(* Logix 5000 project; controller MV vendor 1 type 14 code 217 rev 31.11; software revision 31.00; part 16 of 53 *)
(* tags used below, declared in another part *)
   CWD : CHECKWORD_FLAGS;
   Dummy : BOOL;
   MC_B12 : INT[255];   // PX SWITCH Proxy switch flags f ile
   MC_B240 : INT[255];   // CH1 RN PMP Channel 1 return pum p drive flags
   MC_B241 : INT[255];   // CH2 RN PMP Channel 2 return pum p drive flags
   MC_B242 : INT[255];   // CH1 ROUTE Channel 1 route requ est flags
   MC_B243 : INT[255];   // CH2 ROUTE Channel 2 route requ est flags
   MC_B3 : INT[255];   // BINARY
   MC_bit_data_file_address : DINT;
   MC_bit_file_bit_offset : DINT;
   MC_bit_file_word_offset : DINT;
   MC_bit_offset : DINT;
   MC_bit_returned : BOOL;
   MC_CP1 : PlantItem;   // CP1
   MC_CP1_RawOutput : ALIAS FOR RIO_Rack_2:10:O.Data.14;   // MC_CP1
   MC_data_file_value_to_move : DINT;
   MC_from_data_file : DINT;
   MC_from_data_offset : DINT;
   MC_GBYV1 : PlantItem;   // GBYV1
   MC_GBYV1_RawOutput : ALIAS FOR RIO_Rack_2:8:O.Data.31;   // MC_GBYV1
   MC_N10 : INT[255];   // SETTINGS
   MC_N100 : INT[255];   // C1_PLC Channel 1 PLC data
   MC_N101 : INT[255];   // CH1 PC>PLC Channel 1 PC to PLC
   MC_N102 : INT[255];   // CH1 PROG Channel 1 CIP progra m
   MC_N103 : INT[255];   // CH1 ITEMS Chwd.nos.of items to be checked for Chan nel 1
   MC_N104 : INT[255];   // CH1 REPORT Channel 1 CIP report file
   MC_N108 : INT[255];   // CH1 VDATA Channel 1 CIP progra m validation data
   MC_N112 : INT[255];   // FVR DATA Data read from FV ro uting PLC
   MC_N113 : INT[255];   // MVR DATA Data read from MV ro uting PLC
   MC_N114 : INT[255];   // YP DATA
   MC_N120 : INT[255];   // C2 PLC Channel 2 PLC data
   MC_N121 : INT[255];   // CH2 PC>PLC Channel 2 PC to PLC
   MC_N122 : INT[255];   // CH2 PROG Channel 2 CIP progra m
   MC_N123 : INT[255];   // CH2 ITEMS Chwd.nos.of items to be checked for Chan nel 2
   MC_N124 : INT[255];   // CH2 REPORT Channel 2 CIP report file
   MC_N128 : INT[255];   // CH2 VDATA Channel 2 CIP progra m validation data
   MC_N160 : INT[255];   // P40 CHECK
   MC_N161 : INT[255];   // P41 CHECK
   MC_N162 : INT[255];   // P42 CHECK
   MC_N163 : INT[255];   // P43 CHECK
   MC_N164 : INT[255];   // P44 CHECK
   MC_N165 : INT[255];   // P45 CHECK
   MC_N166 : INT[255];   // P46 CHECK
   MC_N167 : INT[255];   // Original N File From SLC, No Description Available
   MC_N20 : INT[255];   // P1 PRESS Control block and da ta for P1 pressure P ID loop
   MC_N200 : INT[255];   // CHK_WORK Plant item fault che cking work area
   MC_N201 : INT[255];   // P1 CHECK CIP program 1 plant item check list
   MC_N202 : INT[255];   // P2 CHECK CIP program 2 plant item check list
   MC_N203 : INT[255];   // P3 CHECK CIP program 3 plant item check list
   MC_N204 : INT[255];   // P4 CHECK CIP program 4 plant item check list
   MC_N205 : INT[255];   // P5 CHECK CIP program 5 plant item check list
   MC_N206 : INT[255];   // P6 CHECK CIP program 6 plant item check list
   MC_N207 : INT[255];   // P7 CHECK CIP program 7 plant item check list
   MC_N208 : INT[255];   // P8 CHECK CIP program 8 plant item check list
   MC_N209 : INT[255];   // P9 CHECK CIP program 9 plant item check list
   MC_N21 : INT[255];   // P1 FLOW Control block and da ta for P1 flowrate P ID loop
   MC_N210 : INT[255];   // P10 CHECK CIP program 10 plant item check list
   MC_N211 : INT[255];   // P11 CHECK CIP program 11 plant item check list
   MC_N212 : INT[255];   // P12 CHECK CIP program 12 plant item check list
   MC_N213 : INT[255];   // P13 CHECK CIP program 13 plant item check list
   MC_N214 : INT[255];   // P14 CHECK CIP program 14 plant item check list
   MC_N215 : INT[255];   // P15 CHECK CIP program 15 plant item check list
   MC_N216 : INT[255];   // P16 CHECK CIP program 16 plant item check list
   MC_N217 : INT[255];   // P17 CHECK CIP program 17 plant item check list
   MC_N218 : INT[255];   // P18 CHECK CIP program 18 plant item check list
   MC_N219 : INT[255];   // P19 CHECK CIP program 19 plant item check list
   MC_N22 : INT[255];   // P2 PRESS Control block and da ta for P2 pressure P ID loop
   MC_N220 : INT[255];   // P20 CHECK CIP program 20 plant item check list
   MC_N221 : INT[255];   // P21 CHECK CIP program 21 plant item check list
   MC_N222 : INT[255];   // P22 CHECK CIP program 22 plant item check list
   MC_N223 : INT[255];   // P23 CHECK CIP program 23 plant item check list
   MC_N224 : INT[255];   // P24 CHECK CIP program 24 plant item check list
   MC_N225 : INT[255];   // P25 CHECK CIP program 25 plant item check list
   MC_N226 : INT[255];   // P26 CHECK CIP program 26 plant item check list
   MC_N227 : INT[255];   // P27 CHECK CIP program 27 plant item check list
   MC_N228 : INT[255];   // P28 CHECK CIP program 28 plant item check list
   MC_N229 : INT[255];   // P29 CHECK CIP program 29 plant item check list
   MC_N23 : INT[255];   // P2 FLOW Control block and da ta for P2 flowrate P ID loop
   MC_N230 : INT[255];   // P30 CHECK CIP program 30 plant item check list
   MC_N231 : INT[255];   // P31 CHECK CIP program 31 plant item check list
   MC_N232 : INT[255];   // P32 CHECK CIP program 32 plant item check list
   MC_N233 : INT[255];   // P33 CHECK CIP program 33 plant item check list
   MC_N234 : INT[255];   // P34 CHECK CIP program 34 plant item check list
   MC_N235 : INT[255];   // P35 CHECK CIP program 35 plant item check list
   MC_N236 : INT[255];   // P36 CHECK CIP program 36 plant item check list
   MC_N237 : INT[255];   // P37 CHECK CIP program 37 plant item check list
   MC_N238 : INT[255];   // P38 CHECK CIP program 38 plant item check list
   MC_N239 : INT[255];   // P39 CHECK CIP program 39 plant item check list
   MC_N245 : INT[255];   // CC_WORK Continuous checking program work area
   MC_N255 : INT[255];   // CHECKWORDS Plant item checkword s
   MC_N7 : INT[255];   // INTEGER
   MC_N80 : INT[255];   // SRV1_PLC Detergent tank 1 ser vice PLC data
   MC_N81 : INT[255];   // SV1_PC Detergent tank 1 ser vice PC to PLC data
   MC_N82 : INT[255];   // SV1 ITEMS Chwd.nos.of items to be checked for DT1 service
   MC_N90 : INT[255];   // SV2_PLC Detergent tank 2 ser vice PLC data
   MC_N91 : INT[255];   // SV2_PC Detergent tank 2 ser vice PC to PLC data
   MC_N92 : INT[255];   // SV2 ITEMS Chwd.nos.of items to be checked for DT2 service
   MC_SP_V12TO17 : PlantItem;   // SP_V12TO17
   MC_SP_V12TO17_RawOutput : ALIAS FOR RIO_Rack_2:10:O.Data.17;   // MC_SP_V12TO17
(* MC_Common, continued *)

ROUTINE MC_Digital_Outputs   (* ladder *)
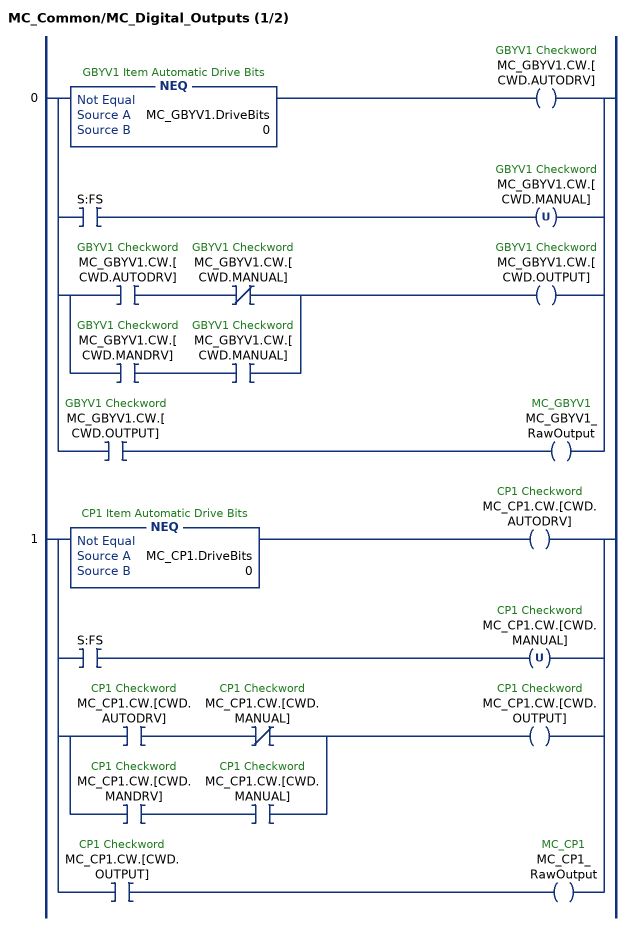
   0: [NEQ(MC_GBYV1.DriveBits,0) OTE(MC_GBYV1.CW.[CWD.AUTODRV]) ,XIC(S:FS) OTU(MC_GBYV1.CW.[CWD.MANUAL]) ,[XIC(MC_GBYV1.CW.[CWD.AUTODRV]) XIO(MC_GBYV1.CW.[CWD.MANUAL]) ,XIC(MC_GBYV1.CW.[CWD.MANDRV]) XIC(MC_GBYV1.CW.[CWD.MANUAL]) ] OTE(MC_GBYV1.CW.[CWD.OUTPUT]) ,XIC(MC_GBYV1.CW.[CWD.OUTPUT]) OTE(MC_GBYV1_RawOutput) ];
   1: [NEQ(MC_CP1.DriveBits,0) OTE(MC_CP1.CW.[CWD.AUTODRV]) ,XIC(S:FS) OTU(MC_CP1.CW.[CWD.MANUAL]) ,[XIC(MC_CP1.CW.[CWD.AUTODRV]) XIO(MC_CP1.CW.[CWD.MANUAL]) ,XIC(MC_CP1.CW.[CWD.MANDRV]) XIC(MC_CP1.CW.[CWD.MANUAL]) ] OTE(MC_CP1.CW.[CWD.OUTPUT]) ,XIC(MC_CP1.CW.[CWD.OUTPUT]) OTE(MC_CP1_RawOutput) ];
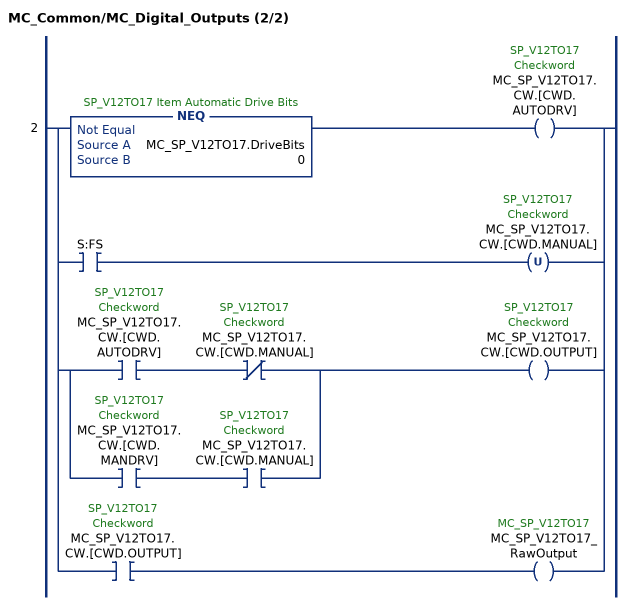
   2: [NEQ(MC_SP_V12TO17.DriveBits,0) OTE(MC_SP_V12TO17.CW.[CWD.AUTODRV]) ,XIC(S:FS) OTU(MC_SP_V12TO17.CW.[CWD.MANUAL]) ,[XIC(MC_SP_V12TO17.CW.[CWD.AUTODRV]) XIO(MC_SP_V12TO17.CW.[CWD.MANUAL]) ,XIC(MC_SP_V12TO17.CW.[CWD.MANDRV]) XIC(MC_SP_V12TO17.CW.[CWD.MANUAL]) ] OTE(MC_SP_V12TO17.CW.[CWD.OUTPUT]) ,XIC(MC_SP_V12TO17.CW.[CWD.OUTPUT]) OTE(MC_SP_V12TO17_RawOutput) ];
END_ROUTINE

ROUTINE MC_Get_NFile_Value   (* ladder *)
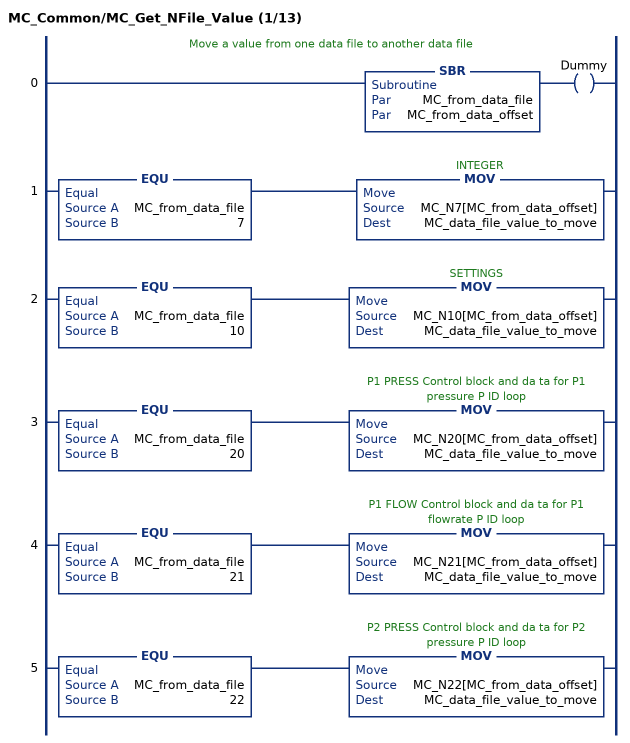
   // Move a value from one data file to another data file
   0: SBR(MC_from_data_file,MC_from_data_offset)OTE(Dummy);
   1: EQU(MC_from_data_file,7)MOV(MC_N7[MC_from_data_offset],MC_data_file_value_to_move);
   2: EQU(MC_from_data_file,10)MOV(MC_N10[MC_from_data_offset],MC_data_file_value_to_move);
   3: EQU(MC_from_data_file,20)MOV(MC_N20[MC_from_data_offset],MC_data_file_value_to_move);
   4: EQU(MC_from_data_file,21)MOV(MC_N21[MC_from_data_offset],MC_data_file_value_to_move);
   5: EQU(MC_from_data_file,22)MOV(MC_N22[MC_from_data_offset],MC_data_file_value_to_move);
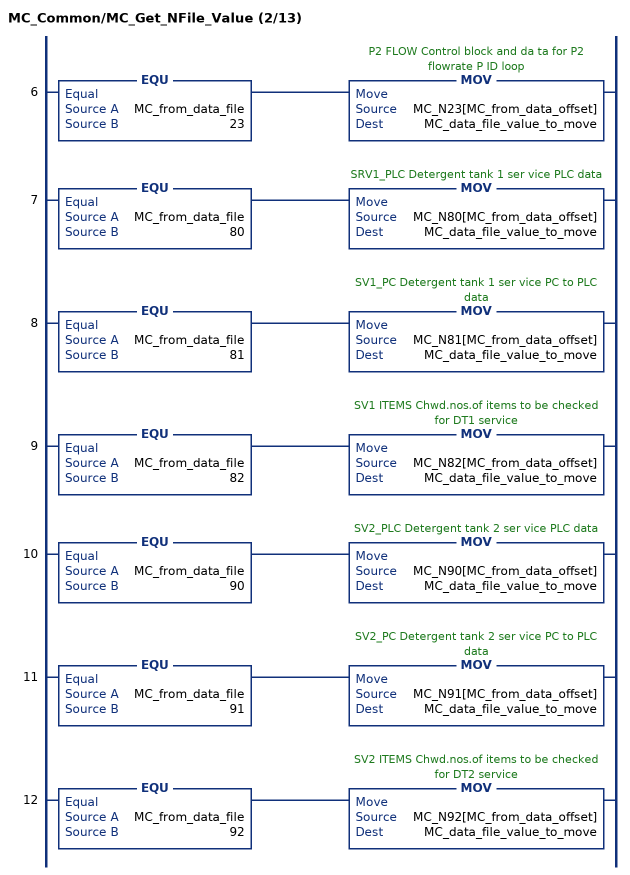
   6: EQU(MC_from_data_file,23)MOV(MC_N23[MC_from_data_offset],MC_data_file_value_to_move);
   7: EQU(MC_from_data_file,80)MOV(MC_N80[MC_from_data_offset],MC_data_file_value_to_move);
   8: EQU(MC_from_data_file,81)MOV(MC_N81[MC_from_data_offset],MC_data_file_value_to_move);
   9: EQU(MC_from_data_file,82)MOV(MC_N82[MC_from_data_offset],MC_data_file_value_to_move);
   10: EQU(MC_from_data_file,90)MOV(MC_N90[MC_from_data_offset],MC_data_file_value_to_move);
   11: EQU(MC_from_data_file,91)MOV(MC_N91[MC_from_data_offset],MC_data_file_value_to_move);
   12: EQU(MC_from_data_file,92)MOV(MC_N92[MC_from_data_offset],MC_data_file_value_to_move);
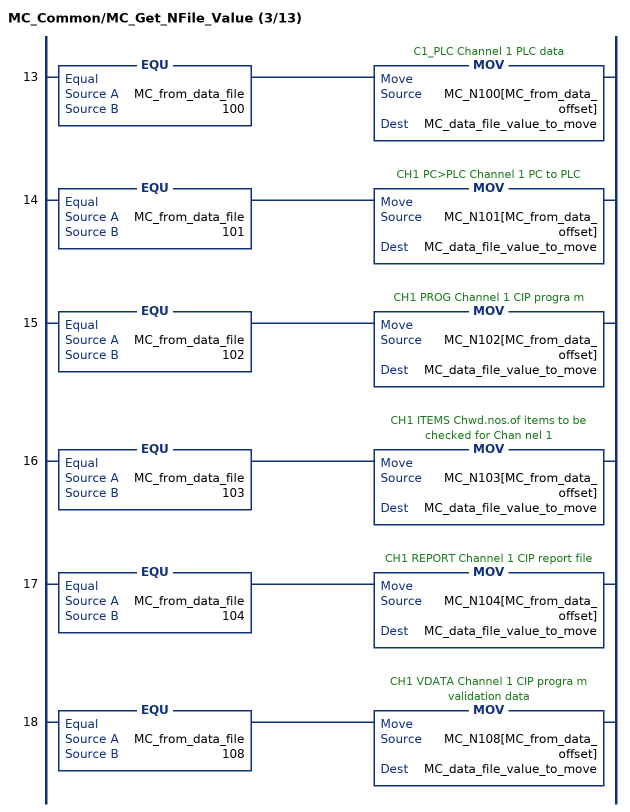
   13: EQU(MC_from_data_file,100)MOV(MC_N100[MC_from_data_offset],MC_data_file_value_to_move);
   14: EQU(MC_from_data_file,101)MOV(MC_N101[MC_from_data_offset],MC_data_file_value_to_move);
   15: EQU(MC_from_data_file,102)MOV(MC_N102[MC_from_data_offset],MC_data_file_value_to_move);
   16: EQU(MC_from_data_file,103)MOV(MC_N103[MC_from_data_offset],MC_data_file_value_to_move);
   17: EQU(MC_from_data_file,104)MOV(MC_N104[MC_from_data_offset],MC_data_file_value_to_move);
   18: EQU(MC_from_data_file,108)MOV(MC_N108[MC_from_data_offset],MC_data_file_value_to_move);
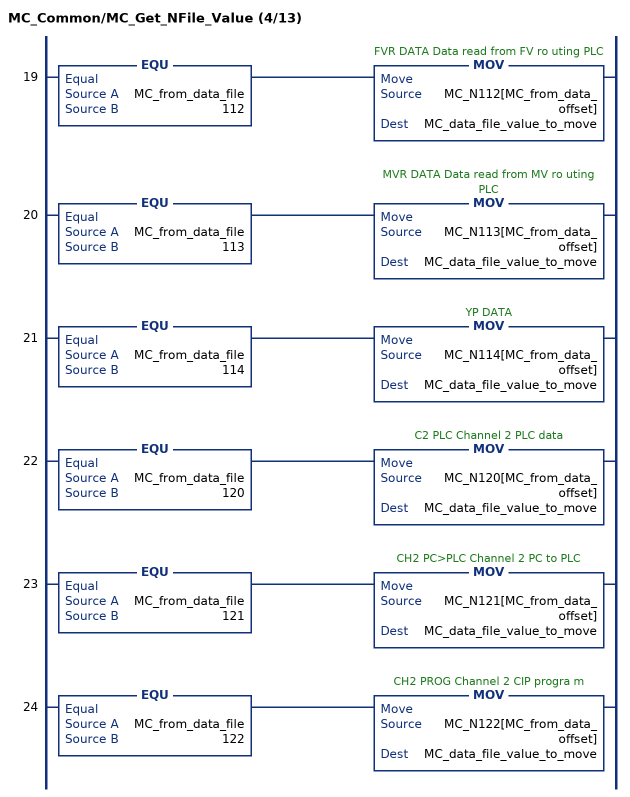
   19: EQU(MC_from_data_file,112)MOV(MC_N112[MC_from_data_offset],MC_data_file_value_to_move);
   20: EQU(MC_from_data_file,113)MOV(MC_N113[MC_from_data_offset],MC_data_file_value_to_move);
   21: EQU(MC_from_data_file,114)MOV(MC_N114[MC_from_data_offset],MC_data_file_value_to_move);
   22: EQU(MC_from_data_file,120)MOV(MC_N120[MC_from_data_offset],MC_data_file_value_to_move);
   23: EQU(MC_from_data_file,121)MOV(MC_N121[MC_from_data_offset],MC_data_file_value_to_move);
   24: EQU(MC_from_data_file,122)MOV(MC_N122[MC_from_data_offset],MC_data_file_value_to_move);
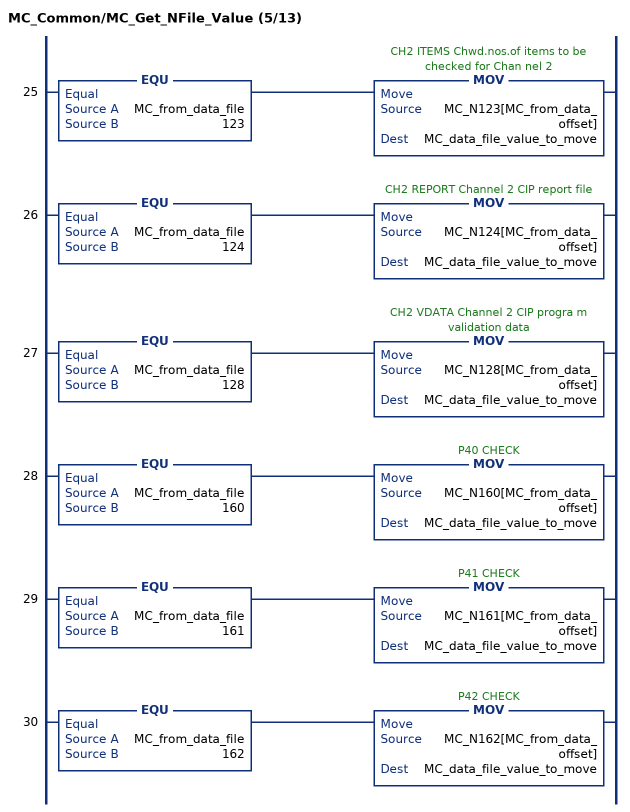
   25: EQU(MC_from_data_file,123)MOV(MC_N123[MC_from_data_offset],MC_data_file_value_to_move);
   26: EQU(MC_from_data_file,124)MOV(MC_N124[MC_from_data_offset],MC_data_file_value_to_move);
   27: EQU(MC_from_data_file,128)MOV(MC_N128[MC_from_data_offset],MC_data_file_value_to_move);
   28: EQU(MC_from_data_file,160)MOV(MC_N160[MC_from_data_offset],MC_data_file_value_to_move);
   29: EQU(MC_from_data_file,161)MOV(MC_N161[MC_from_data_offset],MC_data_file_value_to_move);
   30: EQU(MC_from_data_file,162)MOV(MC_N162[MC_from_data_offset],MC_data_file_value_to_move);
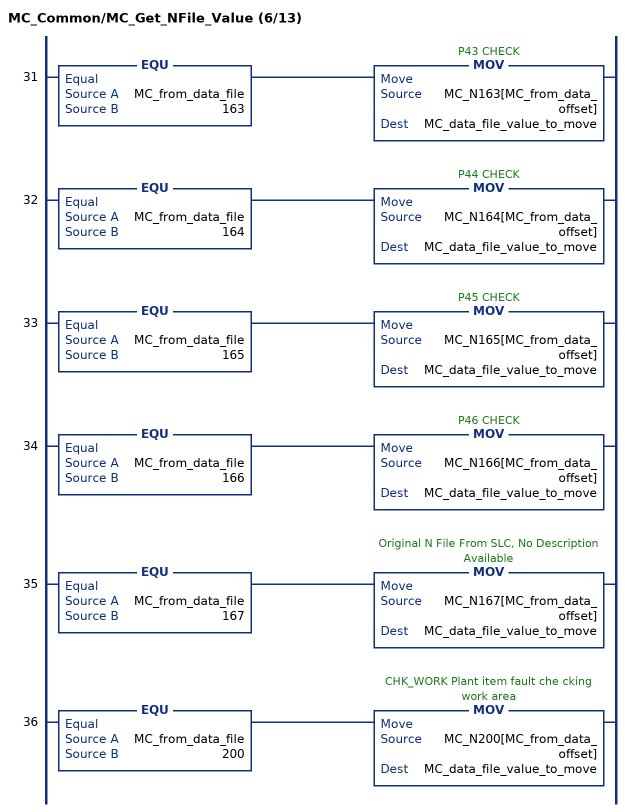
   31: EQU(MC_from_data_file,163)MOV(MC_N163[MC_from_data_offset],MC_data_file_value_to_move);
   32: EQU(MC_from_data_file,164)MOV(MC_N164[MC_from_data_offset],MC_data_file_value_to_move);
   33: EQU(MC_from_data_file,165)MOV(MC_N165[MC_from_data_offset],MC_data_file_value_to_move);
   34: EQU(MC_from_data_file,166)MOV(MC_N166[MC_from_data_offset],MC_data_file_value_to_move);
   35: EQU(MC_from_data_file,167)MOV(MC_N167[MC_from_data_offset],MC_data_file_value_to_move);
   36: EQU(MC_from_data_file,200)MOV(MC_N200[MC_from_data_offset],MC_data_file_value_to_move);
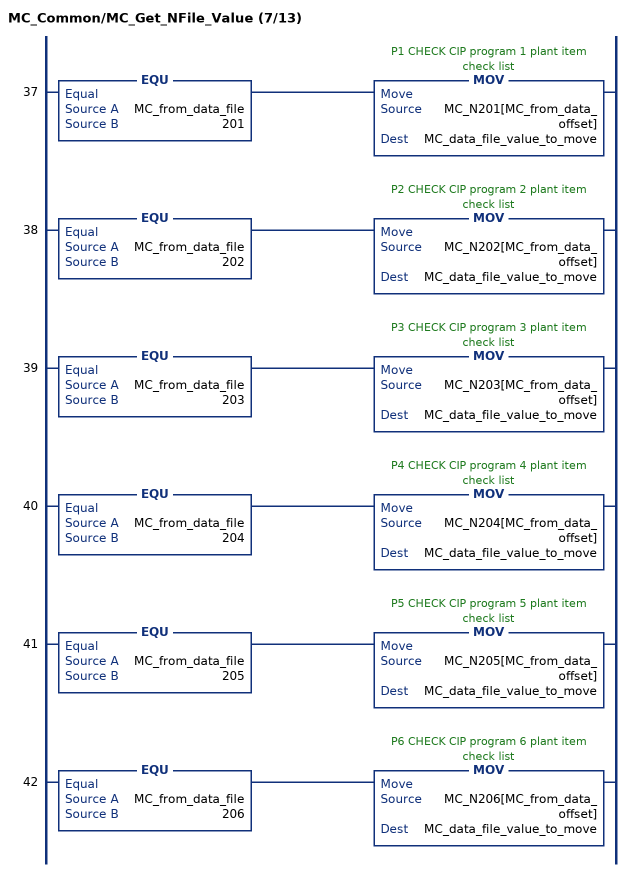
   37: EQU(MC_from_data_file,201)MOV(MC_N201[MC_from_data_offset],MC_data_file_value_to_move);
   38: EQU(MC_from_data_file,202)MOV(MC_N202[MC_from_data_offset],MC_data_file_value_to_move);
   39: EQU(MC_from_data_file,203)MOV(MC_N203[MC_from_data_offset],MC_data_file_value_to_move);
   40: EQU(MC_from_data_file,204)MOV(MC_N204[MC_from_data_offset],MC_data_file_value_to_move);
   41: EQU(MC_from_data_file,205)MOV(MC_N205[MC_from_data_offset],MC_data_file_value_to_move);
   42: EQU(MC_from_data_file,206)MOV(MC_N206[MC_from_data_offset],MC_data_file_value_to_move);
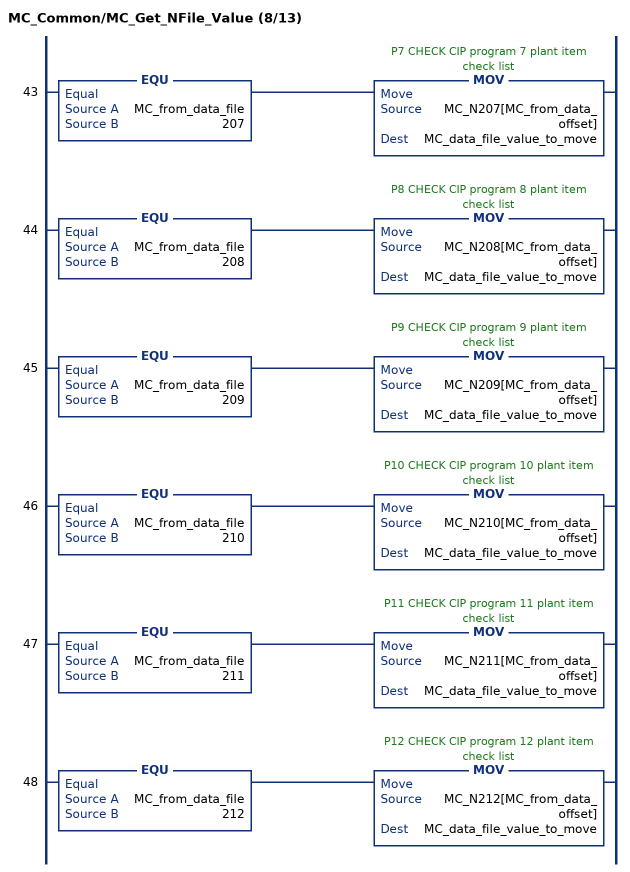
   43: EQU(MC_from_data_file,207)MOV(MC_N207[MC_from_data_offset],MC_data_file_value_to_move);
   44: EQU(MC_from_data_file,208)MOV(MC_N208[MC_from_data_offset],MC_data_file_value_to_move);
   45: EQU(MC_from_data_file,209)MOV(MC_N209[MC_from_data_offset],MC_data_file_value_to_move);
   46: EQU(MC_from_data_file,210)MOV(MC_N210[MC_from_data_offset],MC_data_file_value_to_move);
   47: EQU(MC_from_data_file,211)MOV(MC_N211[MC_from_data_offset],MC_data_file_value_to_move);
   48: EQU(MC_from_data_file,212)MOV(MC_N212[MC_from_data_offset],MC_data_file_value_to_move);
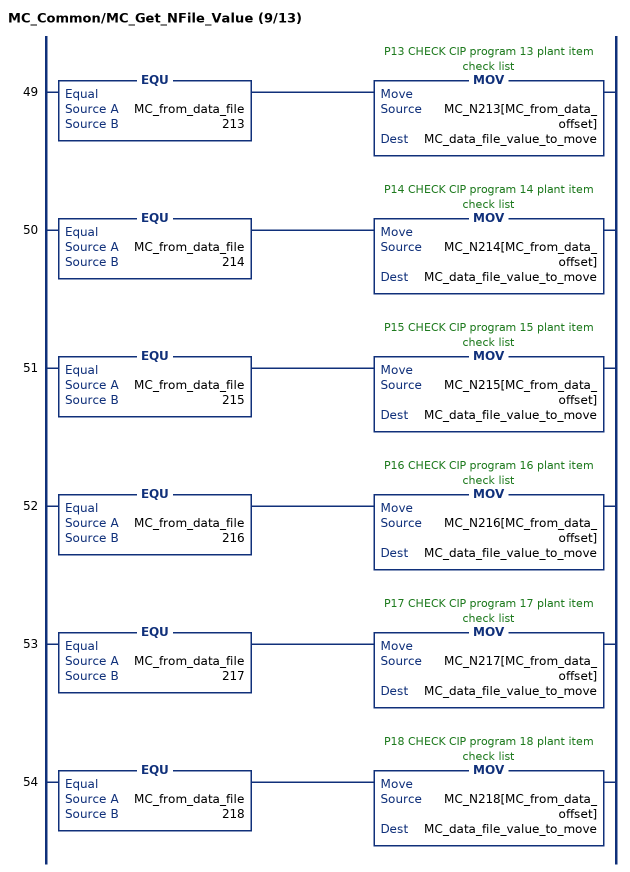
   49: EQU(MC_from_data_file,213)MOV(MC_N213[MC_from_data_offset],MC_data_file_value_to_move);
   50: EQU(MC_from_data_file,214)MOV(MC_N214[MC_from_data_offset],MC_data_file_value_to_move);
   51: EQU(MC_from_data_file,215)MOV(MC_N215[MC_from_data_offset],MC_data_file_value_to_move);
   52: EQU(MC_from_data_file,216)MOV(MC_N216[MC_from_data_offset],MC_data_file_value_to_move);
   53: EQU(MC_from_data_file,217)MOV(MC_N217[MC_from_data_offset],MC_data_file_value_to_move);
   54: EQU(MC_from_data_file,218)MOV(MC_N218[MC_from_data_offset],MC_data_file_value_to_move);
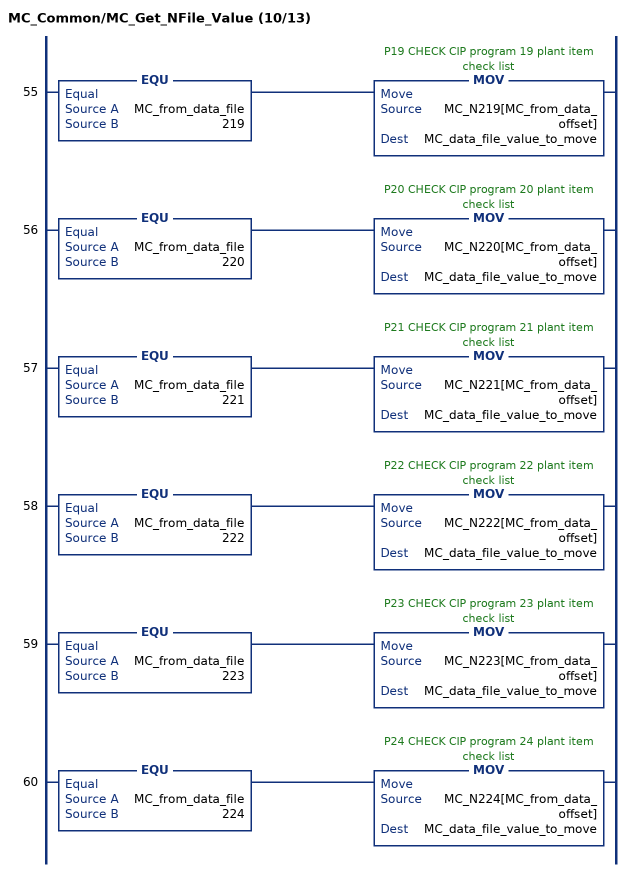
   55: EQU(MC_from_data_file,219)MOV(MC_N219[MC_from_data_offset],MC_data_file_value_to_move);
   56: EQU(MC_from_data_file,220)MOV(MC_N220[MC_from_data_offset],MC_data_file_value_to_move);
   57: EQU(MC_from_data_file,221)MOV(MC_N221[MC_from_data_offset],MC_data_file_value_to_move);
   58: EQU(MC_from_data_file,222)MOV(MC_N222[MC_from_data_offset],MC_data_file_value_to_move);
   59: EQU(MC_from_data_file,223)MOV(MC_N223[MC_from_data_offset],MC_data_file_value_to_move);
   60: EQU(MC_from_data_file,224)MOV(MC_N224[MC_from_data_offset],MC_data_file_value_to_move);
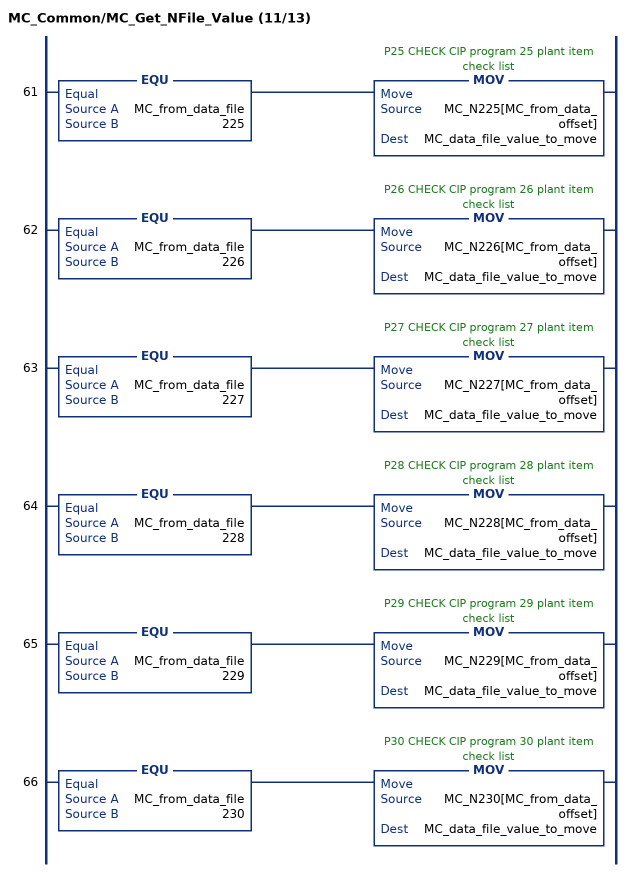
   61: EQU(MC_from_data_file,225)MOV(MC_N225[MC_from_data_offset],MC_data_file_value_to_move);
   62: EQU(MC_from_data_file,226)MOV(MC_N226[MC_from_data_offset],MC_data_file_value_to_move);
   63: EQU(MC_from_data_file,227)MOV(MC_N227[MC_from_data_offset],MC_data_file_value_to_move);
   64: EQU(MC_from_data_file,228)MOV(MC_N228[MC_from_data_offset],MC_data_file_value_to_move);
   65: EQU(MC_from_data_file,229)MOV(MC_N229[MC_from_data_offset],MC_data_file_value_to_move);
   66: EQU(MC_from_data_file,230)MOV(MC_N230[MC_from_data_offset],MC_data_file_value_to_move);
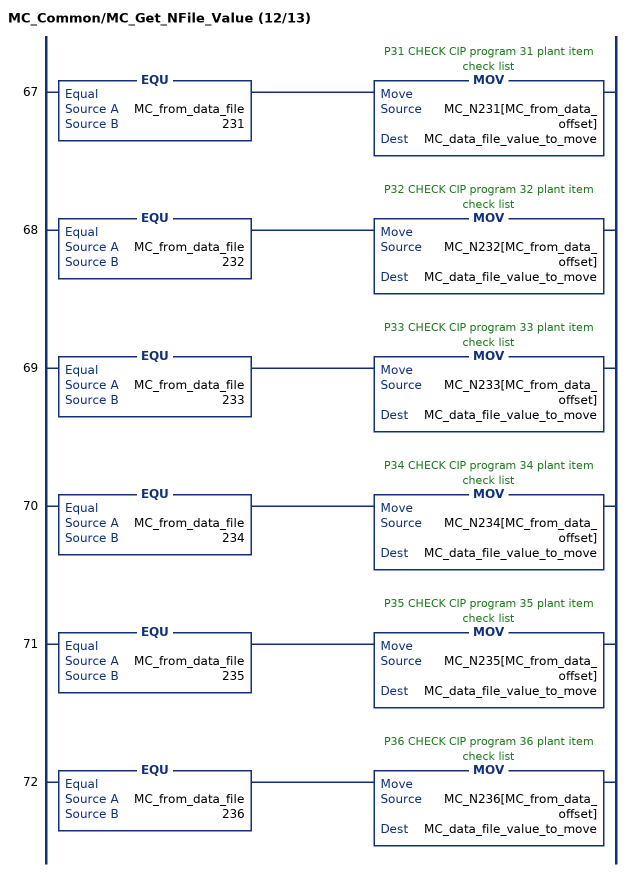
   67: EQU(MC_from_data_file,231)MOV(MC_N231[MC_from_data_offset],MC_data_file_value_to_move);
   68: EQU(MC_from_data_file,232)MOV(MC_N232[MC_from_data_offset],MC_data_file_value_to_move);
   69: EQU(MC_from_data_file,233)MOV(MC_N233[MC_from_data_offset],MC_data_file_value_to_move);
   70: EQU(MC_from_data_file,234)MOV(MC_N234[MC_from_data_offset],MC_data_file_value_to_move);
   71: EQU(MC_from_data_file,235)MOV(MC_N235[MC_from_data_offset],MC_data_file_value_to_move);
   72: EQU(MC_from_data_file,236)MOV(MC_N236[MC_from_data_offset],MC_data_file_value_to_move);
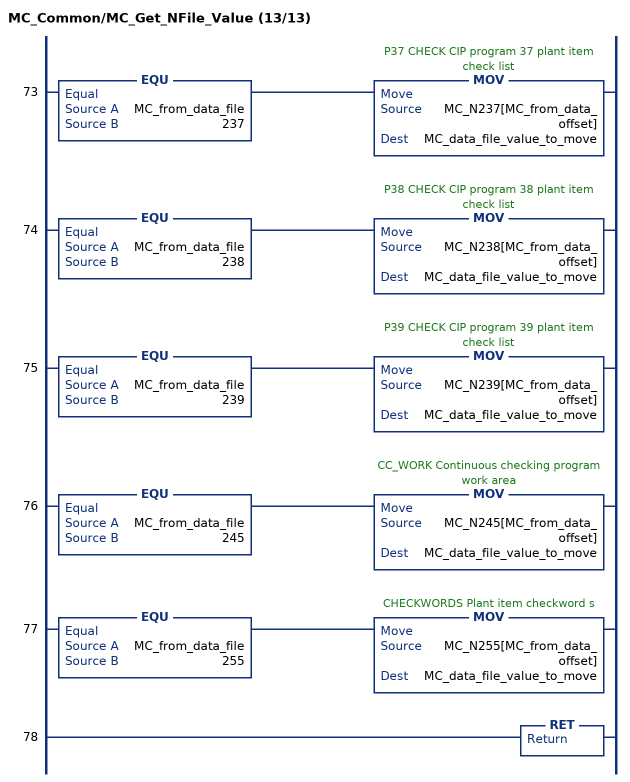
   73: EQU(MC_from_data_file,237)MOV(MC_N237[MC_from_data_offset],MC_data_file_value_to_move);
   74: EQU(MC_from_data_file,238)MOV(MC_N238[MC_from_data_offset],MC_data_file_value_to_move);
   75: EQU(MC_from_data_file,239)MOV(MC_N239[MC_from_data_offset],MC_data_file_value_to_move);
   76: EQU(MC_from_data_file,245)MOV(MC_N245[MC_from_data_offset],MC_data_file_value_to_move);
   77: EQU(MC_from_data_file,255)MOV(MC_N255[MC_from_data_offset],MC_data_file_value_to_move);
   78: RET();
END_ROUTINE

ROUTINE MC_GetBitFile_Value   (* ladder *)
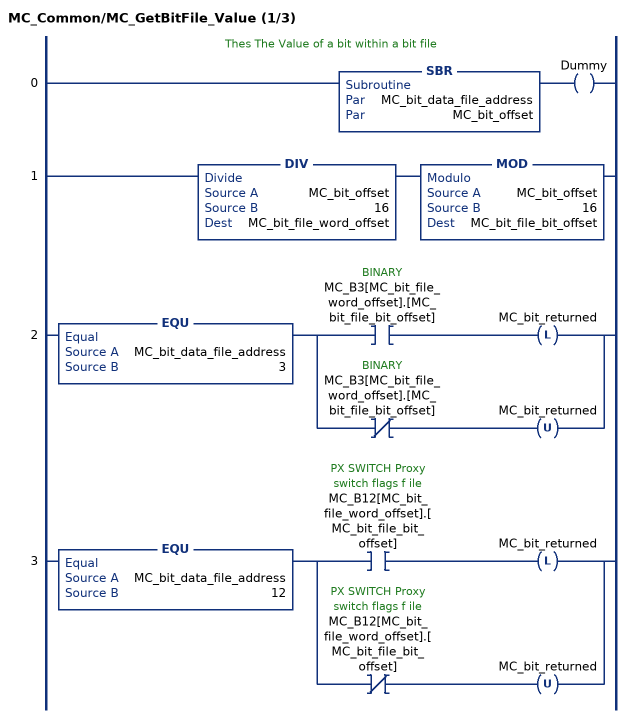
   // Thes The Value of a bit within a bit file
   0: SBR(MC_bit_data_file_address,MC_bit_offset)OTE(Dummy);
   1: DIV(MC_bit_offset,16,MC_bit_file_word_offset)MOD(MC_bit_offset,16,MC_bit_file_bit_offset);
   2: EQU(MC_bit_data_file_address,3)[XIC(MC_B3[MC_bit_file_word_offset].[MC_bit_file_bit_offset]) OTL(MC_bit_returned) ,XIO(MC_B3[MC_bit_file_word_offset].[MC_bit_file_bit_offset]) OTU(MC_bit_returned) ];
   3: EQU(MC_bit_data_file_address,12)[XIC(MC_B12[MC_bit_file_word_offset].[MC_bit_file_bit_offset]) OTL(MC_bit_returned) ,XIO(MC_B12[MC_bit_file_word_offset].[MC_bit_file_bit_offset]) OTU(MC_bit_returned) ];
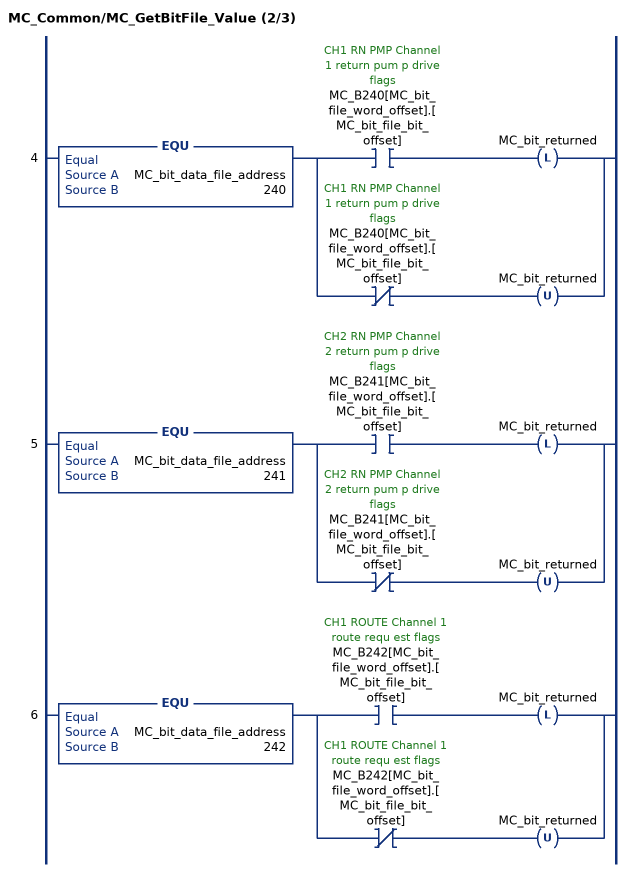
   4: EQU(MC_bit_data_file_address,240)[XIC(MC_B240[MC_bit_file_word_offset].[MC_bit_file_bit_offset]) OTL(MC_bit_returned) ,XIO(MC_B240[MC_bit_file_word_offset].[MC_bit_file_bit_offset]) OTU(MC_bit_returned) ];
   5: EQU(MC_bit_data_file_address,241)[XIC(MC_B241[MC_bit_file_word_offset].[MC_bit_file_bit_offset]) OTL(MC_bit_returned) ,XIO(MC_B241[MC_bit_file_word_offset].[MC_bit_file_bit_offset]) OTU(MC_bit_returned) ];
   6: EQU(MC_bit_data_file_address,242)[XIC(MC_B242[MC_bit_file_word_offset].[MC_bit_file_bit_offset]) OTL(MC_bit_returned) ,XIO(MC_B242[MC_bit_file_word_offset].[MC_bit_file_bit_offset]) OTU(MC_bit_returned) ];
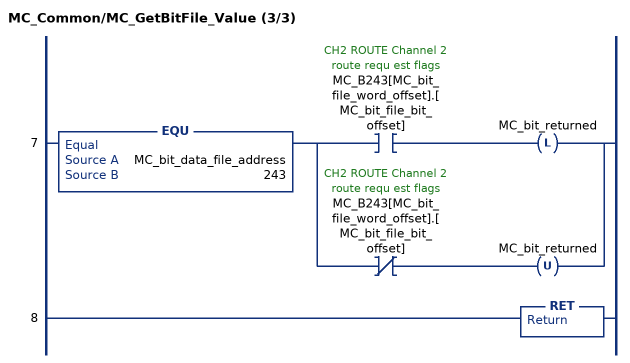
   7: EQU(MC_bit_data_file_address,243)[XIC(MC_B243[MC_bit_file_word_offset].[MC_bit_file_bit_offset]) OTL(MC_bit_returned) ,XIO(MC_B243[MC_bit_file_word_offset].[MC_bit_file_bit_offset]) OTU(MC_bit_returned) ];
   8: RET();
END_ROUTINE
